REGION Network 18: Contrast down
   RUNG wire#powerrail
      Contact( #OS_xNewCapUp )
      Contact( #INO_tTrack.rgtTrackCaps[#AUX_dUpCapIndex].tCap.tDone.xXCutDoneHead )
      { S7_Templates := "SrcType := DInt" } GE_Contact(in1 := #INO_tTrack.rgtTrackCaps[#AUX_dDwCapIndex].tCap.dLength_cmm, in2 := #CONST_DLIMIT_USESNAP_CMM)
      { S7_Templates := "SrcType := DInt" } LE_Contact(in1 := #INO_tTrack.rgtTrackCaps[#AUX_dDwCapIndex].tCap.dLength_cmm, in2 := #tHMW.dMaxPlateLenghtEnableContrast_cmm)
      S_Coil( #tPhases.xContrastDown )
   END_RUNG
   // the same network as SCL:
   IF #OS_xNewCapUp AND #INO_tTrack.rgtTrackCaps[#AUX_dUpCapIndex].tCap.tDone.xXCutDoneHead AND (#INO_tTrack.rgtTrackCaps[#AUX_dDwCapIndex].tCap.dLength_cmm >= #CONST_DLIMIT_USESNAP_CMM) AND (#INO_tTrack.rgtTrackCaps[#AUX_dDwCapIndex].tCap.dLength_cmm <= #tHMW.dMaxPlateLenghtEnableContrast_cmm) THEN
       #tPhases.xContrastDown := TRUE;
   END_IF;
END_REGION

REGION Network 19 (SCL): Calculate contrast activation time
   #TMP_dValue := REAL_TO_DINT(#CONST_DIST_CONTRASTFROMSNAP / #INO_tEnc.rActSpeedValue_cmm_ms + 1500.0);

   IF #TMP_dValue < 0 OR #TMP_dValue>40000 THEN
       #TMP_dValue := 0;
   END_IF;
END_REGION

REGION Network 20: End contrast down
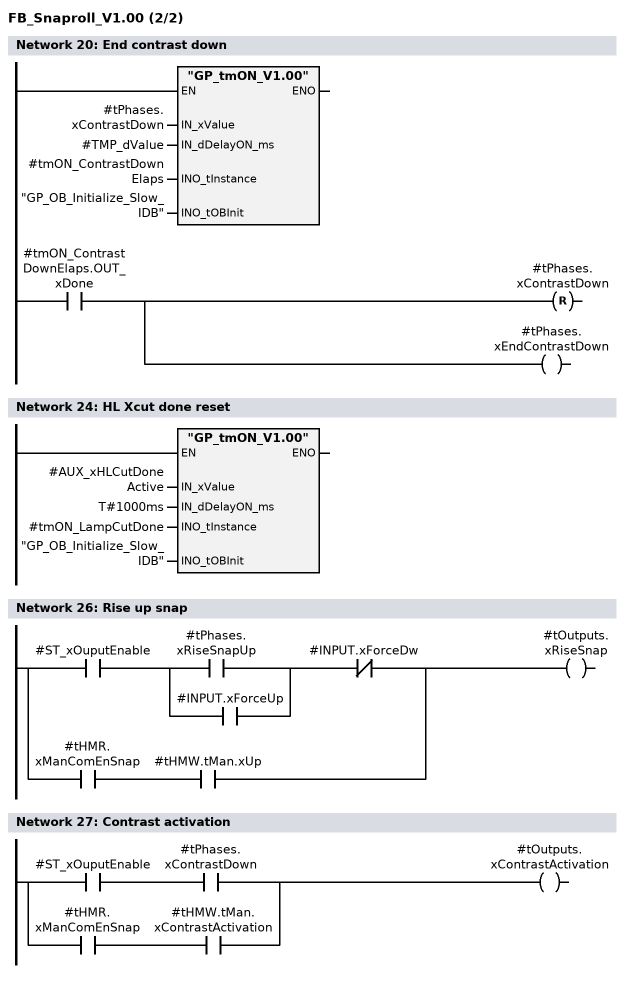
   RUNG wire#powerrail
      "GP_tmON_V1.00"(IN_xValue := #tPhases.xContrastDown, IN_dDelayON_ms := #TMP_dValue, INO_tInstance := #tmON_ContrastDownElaps, INO_tOBInit := "GP_OB_Initialize_Slow_IDB")
   END_RUNG
   RUNG wire#powerrail
      Contact( #tmON_ContrastDownElaps.OUT_xDone )
      wire#w1
      R_Coil( #tPhases.xContrastDown )
   END_RUNG
   RUNG wire#w1
      Coil( #tPhases.xEndContrastDown )
   END_RUNG
   // the same network as SCL:
   "GP_tmON_V1.00"(IN_xValue := #tPhases.xContrastDown,
                   IN_dDelayON_ms := #TMP_dValue,
                   INO_tInstance := #tmON_ContrastDownElaps,
                   INO_tOBInit := "GP_OB_Initialize_Slow_IDB");
   IF #tmON_ContrastDownElaps.OUT_xDone THEN #tPhases.xContrastDown := FALSE; END_IF;
   #tPhases.xEndContrastDown := #tmON_ContrastDownElaps.OUT_xDone;
END_REGION

REGION Network 21 (SCL): ### HMI STATUSES ###
   IF #tOutputs.xRiseSnap THEN
       #tHMR.dStatus := #CONST_DSTATUS_UP;
   ELSIF #ST_xStoppingFaults THEN
       #tHMR.dStatus := #CONST_DSTATUS_ANOMALY;
   ELSE
       #tHMR.dStatus := #CONST_DSTATUS_IDLE;
   END_IF;

   IF #tHMR.xManComEnSnap AND #tHMW.tMan.xUp THEN
       #tHMR.tManCmd.xUp := TRUE;
   ELSE
       #tHMR.tManCmd.xUp := FALSE;
   END_IF;

   IF #tHMR.xManComEnSnap AND #tHMW.tMan.xContrastActivation THEN
       #tHMR.tManCmd.xContrastActivation := TRUE;
   ELSE
       #tHMR.tManCmd.xContrastActivation := FALSE;
   END_IF;
END_REGION

REGION Network 22: ####_OUTPUT_####
END_REGION

REGION Network 23 (SCL): HL Xcut done
   IF #OS_xNewCapUp AND #INO_tTrack.rgtTrackCaps[#AUX_dUpCapIndex].tCap.tDone.xXCutDoneHead THEN
       FOR #TMP_dIndex := 0 TO "DMAXXHEADS_IND" DO
           #tOutputs.rgxHLCutDoneXC[#TMP_dIndex] := #INO_tTrack.rgtTrackCaps[#AUX_dUpCapIndex].tCap.tDone.rgxXCutDoneHead[#TMP_dIndex];
       END_FOR;
       #AUX_xHLCutDoneActive := true;
   END_IF;
END_REGION

REGION Network 24: HL Xcut done reset
   RUNG wire#powerrail
      "GP_tmON_V1.00"(IN_xValue := #AUX_xHLCutDoneActive, IN_dDelayON_ms := T#1000ms, INO_tInstance := #tmON_LampCutDone, INO_tOBInit := "GP_OB_Initialize_Slow_IDB")
   END_RUNG
   // the same network as SCL:
   "GP_tmON_V1.00"(IN_xValue := #AUX_xHLCutDoneActive,
                   IN_dDelayON_ms := T#1000ms,
                   INO_tInstance := #tmON_LampCutDone,
                   INO_tOBInit := "GP_OB_Initialize_Slow_IDB");
END_REGION

REGION Network 25 (SCL): HL Xcut done reset
   IF #tmON_LampCutDone.OUT_xDone THEN
       #AUX_xHLCutDoneActive := false;
       FOR #TMP_dIndex := 0 TO "DMAXXHEADS_IND" DO
           #tOutputs.rgxHLCutDoneXC[#TMP_dIndex] := false;
       END_FOR;
   END_IF;
END_REGION

REGION Network 26: Rise up snap
   RUNG wire#powerrail
      Contact( #ST_xOuputEnable )
      wire#w1
      Contact( #tPhases.xRiseSnapUp )
      wire#w2
      I_Contact( #INPUT.xForceDw )
      wire#w3
      Coil( #tOutputs.xRiseSnap )
   END_RUNG
   RUNG wire#w1
      Contact( #INPUT.xForceUp )
   END_RUNG wire#w2
   RUNG wire#powerrail
      Contact( #tHMR.xManComEnSnap )
      Contact( #tHMW.tMan.xUp )
   END_RUNG wire#w3
   // the same network as SCL:
   #tOutputs.xRiseSnap := (#ST_xOuputEnable AND (#tPhases.xRiseSnapUp OR #INPUT.xForceUp) AND NOT #INPUT.xForceDw) OR (#tHMR.xManComEnSnap AND #tHMW.tMan.xUp);
END_REGION

REGION Network 27: Contrast activation
   RUNG wire#powerrail
      Contact( #ST_xOuputEnable )
      Contact( #tPhases.xContrastDown )
      wire#w1
      Coil( #tOutputs.xContrastActivation )
   END_RUNG
   RUNG wire#powerrail
      Contact( #tHMR.xManComEnSnap )
      Contact( #tHMW.tMan.xContrastActivation )
   END_RUNG wire#w1
   // the same network as SCL:
   #tOutputs.xContrastActivation := (#ST_xOuputEnable AND #tPhases.xContrastDown) OR (#tHMR.xManComEnSnap AND #tHMW.tMan.xContrastActivation);
END_REGION
END_FUNCTION_BLOCK

// folder: 03_Programs_Logics/MCC1200/12_Markers

FUNCTION_BLOCK "FB_Markers_V1.00"   // FB11, LAD
TITLE = Markers bridge V1.00
{ S7_Optimized_Access := 'TRUE' }
VERSION : 0.1
   VAR_INPUT
      IN_xStandardFBCall : Bool;   // FB work modality: Standard call from OB slow
      IN_xCycleON : Bool;   // Cycle ON
      IN_xGeneralReset : Bool;   // General reset
      IN_xResetAlarms : Bool;   // Reset alarms
      IN_xFaultsEnabled : Bool;   // Faults enabled
      IN_tID : Conn_Any;   // Connection ID
      IN_tNewMissionData : "UDT_Marker_Mission_Data";
      IN_tIDeviceData : "UDT_Marker_IDeviceFromBridge";   // IDeviceData from bridge
      IN_dGlassBreakMachineIndex : DInt;   // Glass break machine index
   END_VAR
   VAR_OUTPUT
      OUT_tIDeviceData : "UDT_Marker_IDeviceToBridge";   // IDeviceData to bridge
   END_VAR
   VAR_IN_OUT
      INO_xCallAddTank : Bool;   // FB work modality: Add mission to tank
      INO_tEnc : "UDT_Encoder";   // Encoder data
      INO_tRibbon : "UDT_RibbonData";   // Ribbon data
   END_VAR
   VAR RETAIN
      tHMW : Struct   // HMI Write data
         dSpare : DInt;
      END_STRUCT;
      tHMR : Struct   // HMI Read data
         dSpare : DInt;
      END_STRUCT;
   END_VAR
   VAR
      tALM : Struct   // HMI Alarms
         tS : Struct   // Stopping faults
            xTOutSendData : Bool;   // Timeout send data to bridge
            xSpare_1 : Bool;
            xSpare_2 : Bool;
            xSpare_3 : Bool;
            xSpare_4 : Bool;
            xSpare_5 : Bool;
            xSpare_6 : Bool;
            xSpare_7 : Bool;
            xSpare_8 : Bool;
            xSpare_9 : Bool;
            xSpare_10 : Bool;
            xSpare_11 : Bool;
            xSpare_12 : Bool;
            xSpare_13 : Bool;
            xSpare_14 : Bool;
            xSpare_15 : Bool;
            xSpare_16 : Bool;
            xSpare_17 : Bool;
            xSpare_18 : Bool;
            xSpare_19 : Bool;
            xSpare_20 : Bool;
            xSpare_21 : Bool;
            xSpare_22 : Bool;
            xSpare_23 : Bool;
            xSpare_24 : Bool;
            xSpare_25 : Bool;
            xSpare_26 : Bool;
            xSpare_27 : Bool;
            xSpare_28 : Bool;
            xSpare_29 : Bool;
            xSpare_30 : Bool;
            xSpare_31 : Bool;
         END_STRUCT;
         tF : Struct   // Faults
            xSpare_0 : Bool;
            xSpare_1 : Bool;
            xSpare_2 : Bool;
            xSpare_3 : Bool;
            xSpare_4 : Bool;
            xSpare_5 : Bool;
            xSpare_6 : Bool;
            xSpare_7 : Bool;
            xSpare_8 : Bool;
            xSpare_9 : Bool;
            xSpare_10 : Bool;
            xSpare_11 : Bool;
            xSpare_12 : Bool;
            xSpare_13 : Bool;
            xSpare_14 : Bool;
            xSpare_15 : Bool;
            xSpare_16 : Bool;
            xSpare_17 : Bool;
            xSpare_18 : Bool;
            xSpare_19 : Bool;
            xSpare_20 : Bool;
            xSpare_21 : Bool;
            xSpare_22 : Bool;
            xSpare_23 : Bool;
            xSpare_24 : Bool;
            xSpare_25 : Bool;
            xSpare_26 : Bool;
            xSpare_27 : Bool;
            xSpare_28 : Bool;
            xSpare_29 : Bool;
            xSpare_30 : Bool;
            xSpare_31 : Bool;
         END_STRUCT;
         tW : Struct   // Warnings
            xSpare_0 : Bool;
            xSpare_1 : Bool;
            xSpare_2 : Bool;
            xSpare_3 : Bool;
            xSpare_4 : Bool;
            xSpare_5 : Bool;
            xSpare_6 : Bool;
            xSpare_7 : Bool;
            xSpare_8 : Bool;
            xSpare_9 : Bool;
            xSpare_10 : Bool;
            xSpare_11 : Bool;
            xSpare_12 : Bool;
            xSpare_13 : Bool;
            xSpare_14 : Bool;
            xSpare_15 : Bool;
            xSpare_16 : Bool;
            xSpare_17 : Bool;
            xSpare_18 : Bool;
            xSpare_19 : Bool;
            xSpare_20 : Bool;
            xSpare_21 : Bool;
            xSpare_22 : Bool;
            xSpare_23 : Bool;
            xSpare_24 : Bool;
            xSpare_25 : Bool;
            xSpare_26 : Bool;
            xSpare_27 : Bool;
            xSpare_28 : Bool;
            xSpare_29 : Bool;
            xSpare_30 : Bool;
            xSpare_31 : Bool;
         END_STRUCT;
      END_STRUCT;
      ST_xPhaseInProgress : Bool;   // Phases are in progress
      ST_xPhaseInProgressNetwork : Bool;   // Phase are in progress network
      ST_xStoppingFaults : Bool;   // Stopping faults
      ST_xFaults : Bool;   // Faults
      ST_xWarnings : Bool;   // Warnings
      ST_xOutputEnabled : Bool;   // Output enabled
      ST_xGlassBreak : Bool;   // Glass break under bridge
      tPhases : Struct   // Phases
         xSpare0 : Bool;
         xSpare1 : Bool;
         xSpare2 : Bool;
         xSpare3 : Bool;
         xSpare4 : Bool;
         xSpare5 : Bool;
         xSpare6 : Bool;
         xSpare7 : Bool;
         xSpare8 : Bool;
         xSpare9 : Bool;
         xSpare10 : Bool;
         xSpare11 : Bool;
         xSpare12 : Bool;
         xSpare13 : Bool;
         xSpare14 : Bool;
         xSpare15 : Bool;
         xSpare16 : Bool;
         xSpare17 : Bool;
         xSpare18 : Bool;
         xSpare19 : Bool;
         xSpare20 : Bool;
         xSpare21 : Bool;
         xSpare22 : Bool;
         xSpare23 : Bool;
         xSpare24 : Bool;
         xSpare25 : Bool;
         xSpare26 : Bool;
         xSpare27 : Bool;
         xSpare28 : Bool;
         xSpare29 : Bool;
         xSpare30 : Bool;
         xSpare31 : Bool;
      END_STRUCT;
      tPhasesNetwork : Struct
         xSendMissionInProgr : Bool;   // Send mission data in progress
         xEndSendMissionInProgr : Bool;   // End send mission in progress
         xSendSyncroInProgr : Bool;   // Send syncro in progress
         xEndSendSyncroInProgr : Bool;   // End send syncro in progress
         xSpare4 : Bool;
         xSpare5 : Bool;
         xSpare6 : Bool;
         xSpare7 : Bool;
         xSpare8 : Bool;
         xSpare9 : Bool;
         xSpare10 : Bool;
         xSpare11 : Bool;
         xSpare12 : Bool;
         xSpare13 : Bool;
         xSpare14 : Bool;
         xSpare15 : Bool;
         xSpare16 : Bool;
         xSpare17 : Bool;
         xSpare18 : Bool;
         xSpare19 : Bool;
         xSpare20 : Bool;
         xSpare21 : Bool;
         xSpare22 : Bool;
         xSpare23 : Bool;
         xSpare24 : Bool;
         xSpare25 : Bool;
         xSpare26 : Bool;
         xSpare27 : Bool;
         xSpare28 : Bool;
         xSpare29 : Bool;
         xSpare30 : Bool;
         xSpare31 : Bool;
      END_STRUCT;
      FB_BSEND : BSEND;   // BSend instance
      AUX_tSendDataToBridge : Struct   // Send data to bridge
         tSyncroData : Struct
            dMissionID : DInt;   // Mission Identifier
            dSynchroValue_cmm : DInt;   // Counter value in the last synchro [mm/100]
            dSynchroID : DInt;   // ID of the synchro
            xSpare : Array[0..15] of Bool;
            dSpare : Array[0..9] of DInt;
            iSpare : Int;
         END_STRUCT;
         tMissionData : Struct
            dNumberOfMission : Int;   // Number of mission in packet
            rgtMission : Array[0.."DMAXMARKERMISSIONSEND"] of "UDT_Marker_Mission_Data";   // Missions
         END_STRUCT;
      END_STRUCT;
      ST_xRetrySendMission : Bool;   // Retry send mission
      ST_xRetrySendSyncro : Bool;   // Retry send syncro
      dMissionRecOnTank : DInt;   // Number of received mission on tank
      rgtMissionRecTank : Array[0.."DMAXMARKERMISSIONONTANK"] of "UDT_Marker_Mission_Data";   // Mission tank
   END_VAR
   VAR_TEMP
      TMP_dValue : DInt;
      TMP_dwValue : DWord;
      TMP_iReturn : Int;
      TMP_xCompileMissionData : Bool;
      TMP_dIndex : DInt;
      TMP_wPackLength : Word;
      TMP_xRetrySendMissionWithNewMission : Bool;
      TMP_xRetrySendSyncroWithNewSyncro : Bool;
      TMP_xCompileSyncroData : Bool;
      TMP_xNewCapAvailable : Bool;
   END_VAR
BEGIN

REGION Network 1: ####_CONSTANTS_####
END_REGION

REGION Network 2 (SCL): Mission tank add
   IF #INO_xCallAddTank AND NOT(#IN_xStandardFBCall) THEN
       IF #dMissionRecOnTank <= "DMAXMARKERMISSIONONTANK" THEN

           #rgtMissionRecTank[#dMissionRecOnTank] := #IN_tNewMissionData;
           #dMissionRecOnTank := #dMissionRecOnTank + 1;
       END_IF;
       #INO_xCallAddTank := false;
       RETURN;
   END_IF;

   #IN_xStandardFBCall := 0;
END_REGION

REGION Network 3: ####_MATCH_####
END_REGION

REGION Network 4 (SCL): General reset clean
   IF #IN_xGeneralReset THEN

       #TMP_dwValue := 0;

       SCATTER(IN:=#TMP_dwValue,
               OUT=>#tPhases);

       SCATTER(IN:=#TMP_dwValue,
               OUT=>#tPhasesNetwork);


   END_IF;
END_REGION

REGION Network 5: ####_HMI_LOGICS_####
END_REGION

REGION Network 6 (SCL): List of HMI logics
END_REGION

REGION Network 7: ####_ALARMS_####
END_REGION

REGION Network 8 (SCL): Reset alarms
   IF #IN_xResetAlarms THEN

       #TMP_dwValue := 0;

       SCATTER(IN:=#TMP_dwValue,
               OUT=>#tALM.tF);

       SCATTER(IN:=#TMP_dwValue,
               OUT=>#tALM.tS);

       SCATTER(IN:=#TMP_dwValue,
               OUT=>#tALM.tW);

   END_IF;
END_REGION

REGION Network 9: ####_STATUSES_####
END_REGION

REGION Network 10 (SCL): Calculate alarm statuses
   GATHER(IN:=#tALM.tS,
          OUT=>#TMP_dwValue);

   IF #TMP_dwValue <> 0 THEN
       #ST_xStoppingFaults := TRUE;
   ELSE
       #ST_xStoppingFaults := FALSE;
   END_IF;

   GATHER(IN:=#tALM.tF,
          OUT=>#TMP_dwValue);

   IF #TMP_dwValue <> 0 THEN
       #ST_xFaults := TRUE;
   ELSE
       #ST_xFaults := FALSE;
   END_IF;

   GATHER(IN:=#tALM.tW,
          OUT=>#TMP_dwValue);

   IF #TMP_dwValue <> 0 THEN
       #ST_xWarnings := TRUE;
   ELSE
       #ST_xWarnings := FALSE;
   END_IF;
END_REGION

REGION Network 11 (SCL): Retrieve glass break
   #INO_tRibbon.rgtGlassBreakRequest[#IN_dGlassBreakMachineIndex].IN_dDistanceSnaproll_cmm := #IN_tIDeviceData.rgdDistanceFromSnaproll_cmm[0];
   #INO_tRibbon.rgtGlassBreakRequest[#IN_dGlassBreakMachineIndex].IN_dDownstreamOffset_cmm := 150000;
   #INO_tRibbon.rgtGlassBreakRequest[#IN_dGlassBreakMachineIndex].IN_dUpstreamOffset_cmm := 0;

   IF #INO_tRibbon.rgtGlassBreakRequest[#IN_dGlassBreakMachineIndex].OUT_xDataReady THEN
       #ST_xGlassBreak := #INO_tRibbon.rgtGlassBreakRequest[#IN_dGlassBreakMachineIndex].OUT_xGlassBreak;
   END_IF;

   IF #INO_tRibbon.rgtGlassBreakRequest[#IN_dGlassBreakMachineIndex].OUT_xDataReady OR NOT #INO_tRibbon.rgtGlassBreakRequest[#IN_dGlassBreakMachineIndex].IN_xRequestGlassBreak THEN
       #INO_tRibbon.rgtGlassBreakRequest[#IN_dGlassBreakMachineIndex].OUT_xDataReady := FALSE;
       #INO_tRibbon.rgtGlassBreakRequest[#IN_dGlassBreakMachineIndex].IN_xRequestGlassBreak := TRUE;
   END_IF;
END_REGION

REGION Network 12: ####_PHASES_&_LOGICS_####
END_REGION

REGION Network 13 (SCL): Send mission in progress
   IF NOT #ST_xPhaseInProgressNetwork AND ((#dMissionRecOnTank>0 AND NOT #INO_xCallAddTank) OR #ST_xRetrySendMission) THEN

       IF NOT (#ST_xRetrySendMission) THEN
           #TMP_dValue := #dMissionRecOnTank;
           IF #TMP_dValue > "DMAXMARKERMISSIONSEND" THEN
               #TMP_dValue := "DMAXMARKERMISSIONSEND"+1;
           END_IF;

           FOR #TMP_dIndex := 0 TO "DMAXMARKERMISSIONSEND" DO
               #AUX_tSendDataToBridge.tMissionData.rgtMission[#TMP_dIndex].dPlateID := 0;
               #AUX_tSendDataToBridge.tMissionData.rgtMission[#TMP_dIndex].dMissionID := 0;
               #AUX_tSendDataToBridge.tMissionData.rgtMission[#TMP_dIndex].dMarkerID := 0;
               #AUX_tSendDataToBridge.tMissionData.rgtMission[#TMP_dIndex].dXPosition_cmm := 0;
               #AUX_tSendDataToBridge.tMissionData.rgtMission[#TMP_dIndex].dYPosition_cmm := 0;
               #AUX_tSendDataToBridge.tMissionData.rgtMission[#TMP_dIndex].dSpotSpace_cmm := 0;
           END_FOR;

           #TMP_iReturn := "GP_BlockMoveStruct"(IN_iCount := DINT_TO_INT(#TMP_dValue),
                                                IN_iDestIndex := 0,
                                                IN_iSourceIndex := 0,
                                                INO_vDestArrayStruct := #AUX_tSendDataToBridge.tMissionData.rgtMission,
                                                INO_vSourceArrayStruct := #rgtMissionRecTank);

           #AUX_tSendDataToBridge.tMissionData.dNumberOfMission := DINT_TO_INT(#TMP_dValue);

           #dMissionRecOnTank := #dMissionRecOnTank - #TMP_dValue;

           #TMP_iReturn := "GP_BlockMoveStruct"(IN_iCount := DINT_TO_INT(#dMissionRecOnTank),
                                                IN_iDestIndex := 0,
                                                IN_iSourceIndex := DINT_TO_INT(#TMP_dValue),
                                                INO_vDestArrayStruct := #rgtMissionRecTank,
                                                INO_vSourceArrayStruct := #rgtMissionRecTank);

           FOR #TMP_dIndex := #dMissionRecOnTank TO "DMAXMARKERMISSIONONTANK" DO
               #rgtMissionRecTank[#TMP_dIndex].dPlateID := 0;
               #rgtMissionRecTank[#TMP_dIndex].dMissionID := 0;
               #rgtMissionRecTank[#TMP_dIndex].dMarkerID := 0;
               #rgtMissionRecTank[#TMP_dIndex].dXPosition_cmm := 0;
               #rgtMissionRecTank[#TMP_dIndex].dYPosition_cmm := 0;
               #rgtMissionRecTank[#TMP_dIndex].dSpotSpace_cmm := 0;
           END_FOR;

           #tPhasesNetwork.xSendMissionInProgr := TRUE;
           #ST_xRetrySendMission := FALSE;
           #AUX_tSendDataToBridge.tSyncroData.dMissionID += 1;
       END_IF;

       IF #ST_xRetrySendMission = TRUE THEN
           #tPhasesNetwork.xSendMissionInProgr := TRUE;
           #ST_xRetrySendMission := FALSE;
       END_IF;

   END_IF;
END_REGION

REGION Network 14 (SCL): Send data to bridge
   IF NOT #ST_xPhaseInProgressNetwork AND (#INO_tEnc.xMeterForMarkers OR #ST_xRetrySendSyncro) THEN

       IF #INO_tEnc.xMeterForMarkers THEN

           #AUX_tSendDataToBridge.tSyncroData.dSynchroID += 1;
           #AUX_tSendDataToBridge.tSyncroData.dSynchroValue_cmm := #INO_tEnc.dLastMeterValue_cmm;        

           #INO_tEnc.xMeterForMarkers := FALSE;
           #ST_xRetrySendSyncro := FALSE;
           #tPhasesNetwork.xSendSyncroInProgr := TRUE;
       END_IF;

       IF #ST_xRetrySendSyncro THEN
           #ST_xRetrySendSyncro := FALSE;
           #tPhasesNetwork.xSendSyncroInProgr := TRUE;
       END_IF;

   END_IF;
END_REGION

REGION Network 15: #### SEND DATA TO MARKER ####
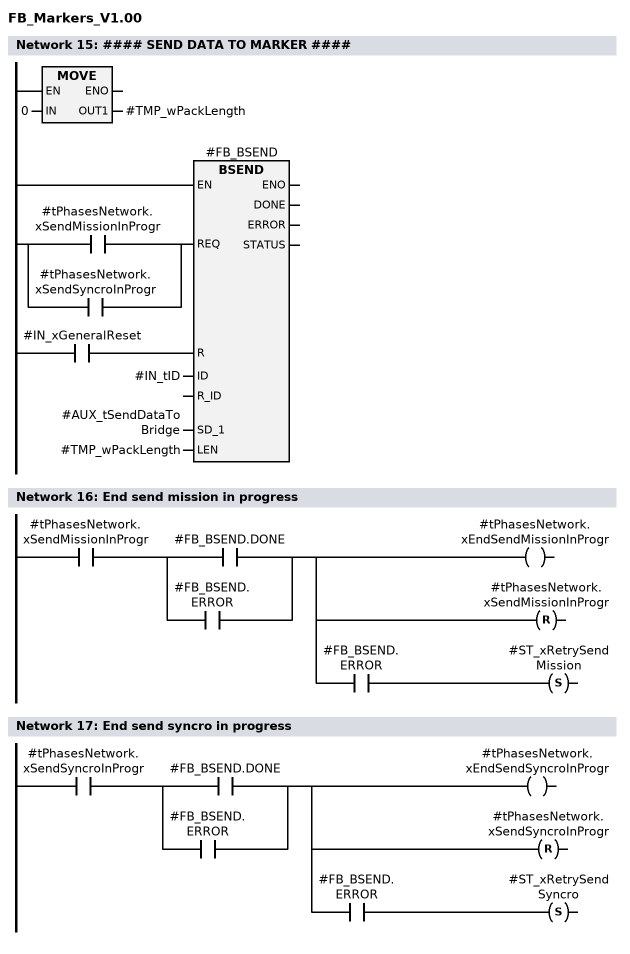
   #TMP_wPackLength := 0;
   #FB_BSEND(REQ := #tPhasesNetwork.xSendMissionInProgr OR #tPhasesNetwork.xSendSyncroInProgr,   // BSEND
             R := #IN_xGeneralReset,
             ID := #IN_tID,
             SD_1 := #AUX_tSendDataToBridge,
             LEN := #TMP_wPackLength);
END_REGION

REGION Network 16: End send mission in progress
   RUNG wire#powerrail
      Contact( #tPhasesNetwork.xSendMissionInProgr )
      wire#w1
      Contact( #FB_BSEND.DONE )
      wire#w2
      Coil( #tPhasesNetwork.xEndSendMissionInProgr )
   END_RUNG
   RUNG wire#w1
      Contact( #FB_BSEND.ERROR )
   END_RUNG wire#w2
   RUNG wire#w2
      R_Coil( #tPhasesNetwork.xSendMissionInProgr )
   END_RUNG
   RUNG wire#w2
      Contact( #FB_BSEND.ERROR )
      S_Coil( #ST_xRetrySendMission )
   END_RUNG
   // the same network as SCL:
   #tPhasesNetwork.xEndSendMissionInProgr := #tPhasesNetwork.xSendMissionInProgr AND (#FB_BSEND.DONE OR #FB_BSEND.ERROR);
   IF #tPhasesNetwork.xEndSendMissionInProgr THEN #tPhasesNetwork.xSendMissionInProgr := FALSE; END_IF;
   IF #tPhasesNetwork.xEndSendMissionInProgr AND #FB_BSEND.ERROR THEN #ST_xRetrySendMission := TRUE; END_IF;
END_REGION

REGION Network 17: End send syncro in progress
   RUNG wire#powerrail
      Contact( #tPhasesNetwork.xSendSyncroInProgr )
      wire#w1
      Contact( #FB_BSEND.DONE )
      wire#w2
      Coil( #tPhasesNetwork.xEndSendSyncroInProgr )
   END_RUNG
   RUNG wire#w1
      Contact( #FB_BSEND.ERROR )
   END_RUNG wire#w2
   RUNG wire#w2
      R_Coil( #tPhasesNetwork.xSendSyncroInProgr )
   END_RUNG
   RUNG wire#w2
      Contact( #FB_BSEND.ERROR )
      S_Coil( #ST_xRetrySendSyncro )
   END_RUNG
   // the same network as SCL:
   #tPhasesNetwork.xEndSendSyncroInProgr := #tPhasesNetwork.xSendSyncroInProgr AND (#FB_BSEND.DONE OR #FB_BSEND.ERROR);
   IF #tPhasesNetwork.xEndSendSyncroInProgr THEN #tPhasesNetwork.xSendSyncroInProgr := FALSE; END_IF;
   IF #tPhasesNetwork.xEndSendSyncroInProgr AND #FB_BSEND.ERROR THEN #ST_xRetrySendSyncro := TRUE; END_IF;
END_REGION

REGION Network 18 (SCL): Calculare phase in progress
   GATHER(IN:=#tPhases,
          OUT=>#TMP_dwValue);

   IF #TMP_dwValue <> 0 THEN
       #ST_xPhaseInProgress := TRUE;
   ELSE
       #ST_xPhaseInProgress := FALSE;
   END_IF;

   GATHER(IN := #tPhasesNetwork,
           OUT => #TMP_dwValue);

   IF  #TMP_dwValue <> 0 THEN
       #ST_xPhaseInProgressNetwork := TRUE;
   ELSE
       #ST_xPhaseInProgressNetwork := FALSE;
   END_IF;
END_REGION

REGION Network 19: ####_OUTPUT_####
END_REGION

REGION Network 20 (SCL): Compile IDevice output
   #OUT_tIDeviceData.xCycleON := #IN_xCycleON;
   #OUT_tIDeviceData.xGlassBreak := #ST_xGlassBreak;
   #OUT_tIDeviceData.xResetAnomaly := #IN_xResetAlarms;
   #OUT_tIDeviceData.xResetBuffers := #IN_xGeneralReset;
   #OUT_tIDeviceData.dSpare2[0] := "DB_Encoder".dActualEncoderCounter_cmm;
END_REGION
END_FUNCTION_BLOCK

// folder: 03_Programs_Logics/MCC1200/13_Z201 comunication

FUNCTION_BLOCK "FB_CommunicationZ300_V1.00"   // FB13, LAD
TITLE = Send data to Z300 V1.00
{ S7_Optimized_Access := 'TRUE' }
VERSION : 0.1
   VAR_INPUT
      IN_dMachineIndex : DInt;   // Tracking machine index
      IN_xCycleON : Bool;   // Cycle ON
      IN_xGeneralReset : Bool;   // General reset
      IN_xResetAlarms : Bool;   // Reset alarms
      IN_dSnapOffset_cmm : DInt;   // Offset on snap [mm/100]
      IN_tID : Conn_Any;   // Connection ID
      tInputs : Struct
         xEmptyingLineArea301 : Bool;   // CS4201 SB
         xStopEmptyingLineArea301 : Bool;   // CS4201 SB
         xResetAnomaly301 : Bool;   // CS4201 SB
         xResetAnomaly302 : Bool;   // CS4201 SB
         xAlarmOFF : Bool;   // CS4201 SB
      END_STRUCT;
      IN_tIDeviceDataIN : "UDT_iDeviceZ301--->Z200";   // IDeviceData from Z300
   END_VAR
   VAR_OUTPUT
      OUT : "UDT_iDevice_MCC1201<---Mcc1200_OUT";
   END_VAR
   VAR_IN_OUT
      INO_tTrack : "UDT_CapData_Tracking";   // Tracking plate
      INO_tEncoder : "UDT_Encoder";   // Encoder data
      INO_xDefectBufferFull : Bool;   // Defect buffer full
      INO_tFBAddDefect : "FB_Defects_Add_V1.00";   // Add defect
      INO_tRibbon : "UDT_RibbonData";   // Ribbon data
      INO_tIDeviceDataOUT : "UDT_iDeviceZ301<---Z200_INO";   // IDevice data to Z300
      INO_tMessage : "UDT_RP_AddMessageCont_v2";   // Message buffer
      INO_xMessageAnomaly : Bool;   // Message anomaly bit
      INO_tMergeSend : "UDT_RP_MessageContMerge_v2";   // Merge buffer to send
      INO_tMergeFromZ300 : "UDT_RP_MessageContMerge_v2";   // Merge buffer from Z300
   END_VAR
   VAR RETAIN
      tHMW : Struct   // HMI Write data
         dAccelerationDelay_ms : DInt;   // Acceleration M301 delay [ms] [mm/100] {ms|s|-1|1|O}
      END_STRUCT;
      tHMR : Struct   // HMI Read data
         dSpare : DInt;
      END_STRUCT;
   END_VAR
   VAR
      tALM : Struct   // HMI Alarms
         tS : Struct   // Stopping faults
            xSpare_0 : Bool;
            xSpare_1 : Bool;
            xSpare_2 : Bool;
            xSpare_3 : Bool;
            xSpare_4 : Bool;
            xSpare_5 : Bool;
            xSpare_6 : Bool;
            xSpare_7 : Bool;
            xSpare_8 : Bool;
            xSpare_9 : Bool;
            xSpare_10 : Bool;
            xSpare_11 : Bool;
            xSpare_12 : Bool;
            xSpare_13 : Bool;
            xSpare_14 : Bool;
            xSpare_15 : Bool;
            xSpare_16 : Bool;
            xSpare_17 : Bool;
            xSpare_18 : Bool;
            xSpare_19 : Bool;
            xSpare_20 : Bool;
            xSpare_21 : Bool;
            xSpare_22 : Bool;
            xSpare_23 : Bool;
            xSpare_24 : Bool;
            xSpare_25 : Bool;
            xSpare_26 : Bool;
            xSpare_27 : Bool;
            xSpare_28 : Bool;
            xSpare_29 : Bool;
            xSpare_30 : Bool;
            xSpare_31 : Bool;
         END_STRUCT;
         tF : Struct   // Faults
            xSpare_0 : Bool;
            xSpare_1 : Bool;
            xSpare_2 : Bool;
            xSpare_3 : Bool;
            xSpare_4 : Bool;
            xSpare_5 : Bool;
            xSpare_6 : Bool;
            xSpare_7 : Bool;
            xSpare_8 : Bool;
            xSpare_9 : Bool;
            xSpare_10 : Bool;
            xSpare_11 : Bool;
            xSpare_12 : Bool;
            xSpare_13 : Bool;
            xSpare_14 : Bool;
            xSpare_15 : Bool;
            xSpare_16 : Bool;
            xSpare_17 : Bool;
            xSpare_18 : Bool;
            xSpare_19 : Bool;
            xSpare_20 : Bool;
            xSpare_21 : Bool;
            xSpare_22 : Bool;
            xSpare_23 : Bool;
            xSpare_24 : Bool;
            xSpare_25 : Bool;
            xSpare_26 : Bool;
            xSpare_27 : Bool;
            xSpare_28 : Bool;
            xSpare_29 : Bool;
            xSpare_30 : Bool;
            xSpare_31 : Bool;
         END_STRUCT;
         tW : Struct   // Warnings
            xSpare_0 : Bool;
            xSpare_1 : Bool;
            xSpare_2 : Bool;
            xSpare_3 : Bool;
            xSpare_4 : Bool;
            xSpare_5 : Bool;
            xSpare_6 : Bool;
            xSpare_7 : Bool;
            xSpare_8 : Bool;
            xSpare_9 : Bool;
            xSpare_10 : Bool;
            xSpare_11 : Bool;
            xSpare_12 : Bool;
            xSpare_13 : Bool;
            xSpare_14 : Bool;
            xSpare_15 : Bool;
            xSpare_16 : Bool;
            xSpare_17 : Bool;
            xSpare_18 : Bool;
            xSpare_19 : Bool;
            xSpare_20 : Bool;
            xSpare_21 : Bool;
            xSpare_22 : Bool;
            xSpare_23 : Bool;
            xSpare_24 : Bool;
            xSpare_25 : Bool;
            xSpare_26 : Bool;
            xSpare_27 : Bool;
            xSpare_28 : Bool;
            xSpare_29 : Bool;
            xSpare_30 : Bool;
            xSpare_31 : Bool;
         END_STRUCT;
      END_STRUCT;
      ST_xPhaseInProgressNetworkPlate : Bool;   // Phase are in progress network plate
      ST_xPhaseInProgressNetworkMessage : Bool;   // Phase are in progress network message
      ST_xPhaseInProgress : Bool;   // Phases are in progress
      ST_xSendDataRequestedPlate : Bool;   // Send plate data
      AUX_xXcutDone : Bool;   // Xcut present
      AUX_xValidUpCap : Bool;   // Upstream cap is valid
      AUX_xValidDwCap : Bool;   // Downstream cap is valid
      AUX_dUpCapIndex : DInt;   // Index of the upstream cap
      AUX_dDwCapIndex : DInt;   // Index of the downstream cap
      AUX_tmonRetainBypassSignal : TOF_TIME;   // Retain bypass snap signal for z300
      AUX_tmonRetainSnapSignal : TOF_TIME;   // Retain snap signal for z300
      OSN_xEndSnapSignal : Bool;   // OSN end of snap signal
      OS_xEndSnapSignal : Bool;   // OS end of snap signal
      OS_xNewCapUp : Bool;   // New cap arrived upstream
      OS_xNewCapDw : Bool;   // New cap arrived downstream
      OS_xNewCapFastDropUp : Bool;   // New cap arrived for fast drop
      OS_xNewCap : Bool;   // New cap arrived
      OS_xEndFastDropSignal : Bool;   // OS end fast drop signal
      OS_xNewCapFastDropUp_1 : Bool;   // New cap arrived for fast drop
      ST_xStoppingFaults : Bool;   // Stopping faults
      ST_xFaults : Bool;   // Faults
      ST_xWarnings : Bool;   // Warnings
      ST_xRetrySendPlate : Bool;   // Retry send
      AUX_xGlassBreakInGoing : Bool;
      AUX_xGlassBreak : Bool;
      AUX_xUpIsQuality : Bool;   // Upstream cap is a quality cap
      AUX_xDwIsQuality : Bool;   // Downstream cap is a quality cap
      AUX_dCounterOnBreak_cmm : DInt;
      tPhases : Struct   // Phases
         xRiseSnapUp : Bool;   // Rise snap
         xEndRiseSnapUp : Bool;   // End rise snap
         xSpare2 : Bool;
         xSpare3 : Bool;
         xSpare4 : Bool;
         xSpare5 : Bool;
         xSpare6 : Bool;
         xSpare7 : Bool;
         xSpare8 : Bool;
         xSpare9 : Bool;
         xSpare10 : Bool;
         xSpare11 : Bool;
         xSpare12 : Bool;
         xSpare13 : Bool;
         xSpare14 : Bool;
         xSpare15 : Bool;
         xSpare16 : Bool;
         xSpare17 : Bool;
         xSpare18 : Bool;
         xSpare19 : Bool;
         xSpare20 : Bool;
         xSpare21 : Bool;
         xSpare22 : Bool;
         xSpare23 : Bool;
         xSpare24 : Bool;
         xSpare25 : Bool;
         xSpare26 : Bool;
         xSpare27 : Bool;
         xSpare28 : Bool;
         xSpare29 : Bool;
         xSpare30 : Bool;
         xSpare31 : Bool;
      END_STRUCT;
      tPhasesNetworkMessage : Struct
         xSendMessageInProgr : Bool;   // Send message data in progress
         xEndSendMessageInProgr : Bool;   // End send message in progress
         xSpare2 : Bool;
         xSpare3 : Bool;
         xSpare4 : Bool;
         xSpare5 : Bool;
         xSpare6 : Bool;
         xSpare7 : Bool;
         xSpare8 : Bool;
         xSpare9 : Bool;
         xSpare10 : Bool;
         xSpare11 : Bool;
         xSpare12 : Bool;
         xSpare13 : Bool;
         xSpare14 : Bool;
         xSpare15 : Bool;
         xSpare16 : Bool;
         xSpare17 : Bool;
         xSpare18 : Bool;
         xSpare19 : Bool;
         xSpare20 : Bool;
         xSpare21 : Bool;
         xSpare22 : Bool;
         xSpare23 : Bool;
         xSpare24 : Bool;
         xSpare25 : Bool;
         xSpare26 : Bool;
         xSpare27 : Bool;
         xSpare28 : Bool;
         xSpare29 : Bool;
         xSpare30 : Bool;
         xSpare31 : Bool;
      END_STRUCT;
      tPhasesNetworkPlate : Struct
         xSendPlateInProgr : Bool;   // Send plate data in progress
         xEndSendPlateInProgr : Bool;   // End send plate data in progress
         xSpare2 : Bool;
         xSpare3 : Bool;
         xSpare4 : Bool;
         xSpare5 : Bool;
         xSpare6 : Bool;
         xSpare7 : Bool;
         xSpare8 : Bool;
         xSpare9 : Bool;
         xSpare10 : Bool;
         xSpare11 : Bool;
         xSpare12 : Bool;
         xSpare13 : Bool;
         xSpare14 : Bool;
         xSpare15 : Bool;
         xSpare16 : Bool;
         xSpare17 : Bool;
         xSpare18 : Bool;
         xSpare19 : Bool;
         xSpare20 : Bool;
         xSpare21 : Bool;
         xSpare22 : Bool;
         xSpare23 : Bool;
         xSpare24 : Bool;
         xSpare25 : Bool;
         xSpare26 : Bool;
         xSpare27 : Bool;
         xSpare28 : Bool;
         xSpare29 : Bool;
         xSpare30 : Bool;
         xSpare31 : Bool;
      END_STRUCT;
      FB_BSEND_PLATE : BSEND;   // BSend plate instance
      FB_BSEND_MESSAGE : BSEND;   // BSend message instance
      AUX_tEmptySendDataToZ300 : "UDT_CapData_Z300";   // Empty send data to Z300
      AUX_tSendDataToZ300 : "UDT_CapData_Z300";   // Send data to Z300
      AUX_tReceivedMerge : "UDT_RP_MessageContMerge_v2";   // Merge received
      FB_BRECV_MESSAGE : BRCV;
      AUX_tCapToSend : "UDT_CapData";
      AUX_dLastInsertDefectPos_cmm : DInt;   // Last inserted defect position [mm/100]
      FB_BRECV_IDEV : BRCV;
      FB_BSEND_IDEV : BSEND;   // BSend plate instance
      AUX_tIDeviceDataIN : "UDT_iDeviceZ301--->Z200";   // IDeviceData from Z300
   END_VAR
   VAR_TEMP
      TMP_dValue : DInt;
      TMP_lwValue : LWord;
      TMP_dwValue : DWord;
      TMP_dIndex : DInt;
      TMP_wPackLength : Word;
      TMP_xNewCapAvailable : Bool;
      TMP_rgxWValue : Array[0..15] of Bool;
      TMP_rgxDWValue : Array[0..31] of Bool;
      TMP_wValue : Word;
      TMP_dConvNumPlate : DInt;
      TMP_dConvTotalLength_cmm : DInt;
      TMP_dConvGap_cmm : DInt;
      TMP_dNumMessage : DInt;
      TMP_dPos : DInt;
      TMP_iRet : Int;
      TMP_dSerializePos : DInt;
      TMP_rgbDInt : Array[0..3] of Byte;
      DEBUG_xVal1 : Bool;
      TMP_dTrackTail : DInt;
      TMP_dMexIndex : DInt;
      TMP_xExit : Bool;
      TMP_xCutDone : Bool;
      TMP_xReqDoneMatch : Bool;
      TMP_xGlassBreak : Bool;
      TMP_dEncDef_cmm : DInt;
   END_VAR
   VAR CONSTANT
      CONST_DSTATUS_IDLE : DInt := 1;   // Status idle
      CONST_DSTATUS_UP : DInt := 3;   // Status up
      CONST_DSTATUS_ANOMALY : DInt := 7;   // Status anomaly
      CONST_MINPLATELENGTH_Z300_CMM : DInt := 60000;   // Minimum plate lenght to send to Z300